
       #FB_STATE_TCP_RECONNECTING:
         REGION FB_STATE_TCP_RECONNECTING
           IF #tempTsendcStatus = #TSENDC_EST_OK THEN
             #statErrorAutoCleared := FALSE;
             //Monitor Connection
             #statFBState := #FB_STATE_OPERATING_MONITOR_TCP;
             // Begin MQTT Connection
             #statMqttConnectState := #MQTT_CONNECT_STATE_BUILD_PAKET;
           END_IF;
         END_REGION FB_STATE_TCP_RECONNECTING
       #FB_STATE_DISABLING: // Disabling active
         REGION DISABLING FB
           //  Disabling, e.g. closing connections, etc.
           // When disabling is complete the bit #statDisablingCompleted must be set
           // When MQTT is connected, send disconnect
           IF #statMqttConnectState = #MQTT_CONNECT_STATE_CONNECTED THEN
             IF #statTsendcReq = TRUE THEN
               //Interrupt any existing send jobs
               #statTsendcReq := FALSE;
             ELSE
               // INIT
               #statSendBufferPos := 0;
               //Build fixed Header
               //Message Type
               #statSendBuffer[#statSendBufferPos] := #MQTT_MSG_TYPE_DISCONNECT;
               #statSendBufferPos += 1;
               //Remaining Length (must be O)
               #statSendBuffer[#statSendBufferPos] := #REMAINIG_LEN_0;
               #statSendBufferPos += 1;
               //send request
               #statTsendcLen := #statSendBufferPos;
               #statTsendcReq := TRUE;
               #statMqttConnectState := #MQTT_CONNECT_STATE_DISCONNECTED;
             END_IF;
           ELSE
             //Disable TCP Connection
             #statTsendcReq := FALSE;
             #statTsendcEnable := FALSE;
             #statEnableTimerCommandWatchdog := TRUE;
           END_IF;
           // When TCP connection is closed
           IF #tempTsendcStatus = #TSENDC_DISCONNECTED THEN
             #statEnableTimerCommandWatchdog := FALSE;
             #statDisablingCompleted := TRUE;
           ELSIF #instTimerCommandWatchdog.Q THEN
             #statEnableTimerCommandWatchdog := FALSE;
             #statDisablingCompleted := TRUE;
           END_IF;
         END_REGION DISABLING FB
       ELSE // Undefined state in state machine reached
         #statStatus := #ERR_UNDEFINED_STATE;
         #statErrorUserCleared := TRUE;
     END_CASE;
   END_REGION STATE_MACHINE

   REGION OUTPUTS
     // Write outputs
     IF (#statDisablingCompleted = TRUE) THEN
       // Reset outputs if disabling completed
       #statValid := FALSE;
       #statBusy := FALSE;
       #statError := FALSE;
       #statDone := FALSE;
       #statErrorUserCleared := FALSE;
       #statErrorAutoCleared := FALSE;
       #statStatus := #STATUS_NO_CALL;
       // Reset application specific outputs
       #statRcvMsgStatus := #MSG_DECODE_STATUS_NO_NEW_MSG;
       #statRcvMsgDataLen := 0;
     ELSIF (#statErrorUserCleared = TRUE) AND (#statError = FALSE) THEN
       // Error can only be cleared by user; rising edge at enable input is needed to continue 
       #statValid := FALSE;
       #statBusy := FALSE;
       #statDone := FALSE;
       #statError := TRUE;
       // Write diagnostics
       #diagnostics.status := #statStatus;
       #diagnostics.subfunctionStatus := #statSubfunctionStatus;
       #diagnostics.stateNumber := #statFBErrorState;
       // execution aborted --> set state no processing
       #statTsendcEnable := FALSE; // Terminate Connection, no reason keep it up.
       #statFBState := #FB_STATE_NO_PROCESSING;
       #statMqttConnectState := #MQTT_CONNECT_STATE_NO_PROCESSING;
       #statMqttCommandState := #MQTT_COMMAND_STATE_NO_PROCESSING;
       #statRcvMsgDecodeState := #MSG_DECODE_STATE_NO_PROCESSING;

     ELSIF (#statErrorAutoCleared = TRUE) AND (#statError = FALSE) THEN
       // Error can be reset by FB automatically
       #statValid := FALSE;
       #statBusy := TRUE;
       #statError := TRUE;
       #statDone := FALSE;
       // Write diagnostics
       #diagnostics.status := #statStatus;
       #diagnostics.subfunctionStatus := #statSubfunctionStatus;
       #diagnostics.stateNumber := #statFBErrorState;
       // Handling of autocleared error
       CASE #statStatus OF
           //Just signal error and reset autocleared error afterwards.
         #ERR_MQTT_PAKET_ID_INVALID, #ERR_MQTT_SUBACK_FAILURE, #ERR_MQTT_CONNECT_TIMEOUT,
         #ERR_MQTT_COMMAND_SEND_TIMEOUT, #ERR_MQTT_COMMAND_MULTIPLE_INPUT, #ERR_CNT_EXCEEDS_ARRAY_DIMENSION,
         #ERR_MQTT_COMMAND_PUBLISH_TOPIC_INVALID, #ERR_QOS_INVALID, #ERR_MQTT_COMMAND_SUBSCRIBE_TOPIC_INVALID:
           #statErrorAutoCleared := FALSE;

         ELSE  // Statement section ELSE
           ;
       END_CASE;

     ELSIF (#statErrorAutoCleared = FALSE) AND (#statErrorUserCleared = FALSE) AND (#statError = TRUE) THEN
       // If autocleared error is acknowledged
       #statValid := TRUE;
       #statBusy := TRUE;
       #statError := FALSE;
       #statDone := FALSE;
       //   this line  more detailed status information is used instead of "#STATUS_SUBSEQUENT_CALL"
       CASE #statStatus OF
         #ERR_TCP_RECONNECTING, #ERR_MQTT_CONNECT_TIMEOUT:  // Reconnecting ok, start Mqtt reconnnect
           //set status
           #statStatus := #STATUS_MQTT_CONNECTING;
           //in the following status codes status stays connected. 
         #ERR_MQTT_PAKET_ID_INVALID, #ERR_MQTT_SUBACK_FAILURE, #ERR_MQTT_COMMAND_SEND_TIMEOUT,
         #ERR_MQTT_COMMAND_MULTIPLE_INPUT, #ERR_CNT_EXCEEDS_ARRAY_DIMENSION, #ERR_MQTT_COMMAND_PUBLISH_TOPIC_INVALID,
         #ERR_QOS_INVALID, #ERR_MQTT_COMMAND_SUBSCRIBE_TOPIC_INVALID:
           #statStatus := #STATUS_MQTT_CONNECTED;
         ELSE  // Statement section ELSE
           ;
       END_CASE;
     END_IF;

     // Write static values to outputs
     #valid := #statValid;
     #busy := #statBusy;
     #error := #statError;
     #status := #statStatus;
     //block sets ENO automatically:
     //ENO := TRUE;
     //Write application specific static values to outputs
     #done := #statDone;
     #receivedMsgStatus := #statRcvMsgStatus;
     #receivedMsgDataLen := #statRcvMsgDataLen;
   END_REGION OUTPUTS
END_FUNCTION_BLOCK

// folder: LMQTT/Utilities

FUNCTION "LMQTT_ConvertToUtf8" : Void   // FC6, SCL
TITLE = LMQTT_ConvertToUtf8
{ S7_Optimized_Access := 'TRUE' }
AUTHOR : SIEMENS
FAMILY : LMQTT
VERSION : 1.0
// Function to convert a WCHAR to a UTF-8 conformant byte sequence
   VAR_INPUT
      character : WChar;   // Character that shall be converted to UTF-8
   END_VAR
   VAR_OUTPUT
      convertedUtf8 : DWord;   // UTF-8 conformant byte sequence. B0 stores first Byte, B1 second and B2 third Byte. B3 is not used
      bytesUsed : USInt;   // Amount of Bytes converted. Ranges from 1 to 3.
      error : Bool;   // TRUE: An error occurred during the execution of the FC
      status : Word;   // 16#0000 - 16#7FFF: Status of the FC, 16#8000 - 16#FFFF: Error identification
   END_VAR
   VAR_TEMP
      tempStatus : Word;   // temp value for output 'status'
      tempConvertedUtf8 : DWord;   // temp value for output 'convertedUtf8'
      tempBytesUsed : USInt;   // temp value for output 'bytesUsed'
      tempCharacter : WChar;   // temp value for input 'character'
   END_VAR
   // Ret_Val : No return for this FC - see error and status output
   VAR CONSTANT
      STATUS_NO_ERROR : Word := 16#0000;   // no error status
      STATUS_EXECUTION_FINISHED : Word := 16#0000;   // Execution finished without errors
      ERR_UNDEFINED : Word := 16#8000;   // Error due to an undefined case
      USINT_NULL : USInt := 0;   // Init value with 0
      DWORD_NULL : DWord := 16#0000_0000;   // Init value with 0
      EMPTY_WCHAR : WChar := WCHAR#' ';   // Empty WChar for comparison
      BELOW_7F : Word := 16#007F;   // Upper limit for character if only one Byte used
      BELOW_7FF : Word := 16#07FF;   // Upper limit for character if two Byte used
      BELOW_MAX_FFFF : Word := 16#FFFF;   // Upper limit for character if three Byte used
      BYTE_3F : Byte := 16#3F;   // Conversion Value
      BYTE_80 : Byte := 16#80;   // Conversion Value
      BYTE_C0 : Byte := 16#C0;   // Conversion Value
      BYTE_E0 : Byte := 16#E0;   // Conversion Value
      USINT_ONE : USInt := 1;   // Const Value to assign amount of bytes used
      USINT_TWO : USInt := 2;   // Const Value to assign amount of bytes used
      USINT_THREE : USInt := 3;   // Const Value to assign amount of bytes used
   END_VAR
BEGIN
   REGION BLOCK INFO HEADER
       //=============================================================================
       // SIEMENS AG
       // (c)Copyright 2020
       //-----------------------------------------------------------------------------
       // Library:       LMQTT
       // Tested with:   CPU 1516-3 PN/DP V2.8
       // Engineering:   TIA Portal V16
       // Restrictions:  --
       // Requirements:  --
       // Functionality: Converts a single WChar Character to a valid UTF-8 encoded byte sequence and saves this to a DWord.
       //                The amount of bytes saved is stored in bytesUsed Output.
       //-----------------------------------------------------------------------------
       // Change log table:
       // Version    Date         Expert in charge         Changes applied
       // 03.00.00   01.10.2020   Siemens Online Support   First released version
       //=============================================================================
   END_REGION

   REGION INITIALISATION  
       // Initialize functionality: reset of variables, diagnostics, etc.
       #tempConvertedUtf8 := #DWORD_NULL;
       #tempBytesUsed := #USINT_NULL;
       #tempStatus := #STATUS_NO_ERROR;
       //assign temp value from input:
        #tempCharacter := #character;

   END_REGION

   REGION PROGRAM LOGIC
       // Use this region for application specific code
       IF #tempCharacter = #EMPTY_WCHAR THEN
           //will be only 1 byte occupied
           #tempConvertedUtf8 := WCHAR_TO_DWORD(#tempCharacter);
           #tempBytesUsed := #USINT_ONE;
       ELSIF (WCHAR_TO_WORD(#tempCharacter) <= (#BELOW_7F)) THEN
           //will be only 1 byte occupied
           #tempConvertedUtf8 := WCHAR_TO_DWORD(#tempCharacter);
           #tempBytesUsed := #USINT_ONE;
       ELSIF (WCHAR_TO_WORD(#tempCharacter) <= (#BELOW_7FF)) THEN
           //will be 2 byte occupied
           #tempConvertedUtf8.%B1 := (WCHAR_TO_BYTE(#tempCharacter) AND #BYTE_3F) OR #BYTE_80;
           #tempConvertedUtf8.%B0 := WORD_TO_BYTE(SHR(IN := WCHAR_TO_WORD(#tempCharacter), N := 6)) OR #BYTE_C0;
           #tempBytesUsed := #USINT_TWO;
       ELSIF (WCHAR_TO_WORD(#tempCharacter) <= (#BELOW_MAX_FFFF)) THEN
           //will be 3 byte occupied
           #tempConvertedUtf8.%B2 := (WCHAR_TO_BYTE(#tempCharacter) AND #BYTE_3F) OR #BYTE_80;
           #tempConvertedUtf8.%B1 := (WORD_TO_BYTE(SHR(IN := WCHAR_TO_WORD(#tempCharacter), N := 6)) AND #BYTE_3F) OR #BYTE_80;
           #tempConvertedUtf8.%B0 := WORD_TO_BYTE(SHR(IN := WCHAR_TO_WORD(#tempCharacter), N := 12)) OR #BYTE_E0;
           #tempBytesUsed := #USINT_THREE;
       END_IF;
   END_REGION

   REGION OUTPUTS
       // Write application specific temp values to outputs
       #bytesUsed := #tempBytesUsed;
       #convertedUtf8 := #tempConvertedUtf8;
       // Write error and status
       #error := #tempStatus.%X15;
       #status := #tempStatus;
       // ENO mechanism is not used --> ENO := TRUE;
       ENO := TRUE;
   END_REGION
END_FUNCTION

// folder: LStream

FUNCTION_BLOCK "LStream_JsonDeserializer"   // FB3, SCL
TITLE = LStream_JsonDeserializer / LStream_JsonParser
{ S7_Optimized_Access := 'TRUE' }
AUTHOR : DI_FA_S_SUP_EuC
FAMILY : LStream
VERSION : 1.0
// parses a JSON string provided in the raw paramter  and rebuilds the coinatend bytes into a tree structure / Parses JSON file, with or without seach option
   VAR_INPUT
      execute : Bool;   // Rising edge starts action once
      search : Bool;   // TRUE: Search option is acticve
   END_VAR
   VAR_OUTPUT
      done : Bool;   // TRUE: Commanded functionality has been completed successfully
      busy : Bool;   // TRUE: FB is not finished and new output values can be expected
      error : Bool;   // TRUE: An error occurred during the execution of the FB
      status : Word := 16#7000;   // 16#0000 - 16#7FFF: Status of the FB, 16#8000 - 16#FFFF: Error identification
      resultCount : Int;   // Count of parsed JSON elements
   END_VAR
   VAR_IN_OUT
      tree : Array[*] of "LStream_typeElement";   // JSON tree containing the stored data
      raw : Array[*] of Byte;   // raw JSON data to parse in byte format
   END_VAR
   VAR
      statExecuteOld : Bool;   // Old value of 'execute' input for edge detection
      statDone : Bool;   // Static value for output 'done'
      statBusy : Bool;   // Static value for output 'busy'
      statError : Bool;   // Static value for output 'error'
      statStatus : Word := 16#7000;   // Static value for output 'status'
      statFBState : DInt := 0;   // State in the state machine of the FB
      statCountOfTree : Int;   // Static count of tree fields
      statCountOfRaw : Int;   // Static count of raw fields
      statResultCount : Int;   // Static value of result count
      statRawIndex : Int;   // Static value of raw index
      instWatchdog : IEC_TIMER;   // instance of watchdog timer
      statSearch : Bool;   // TRUE: Only keys provided in tree will be parsed
      statKeyValueFound : Bool;   // TRUE: Key exisits in raw data
      statTreeIndex : Int;   // Static value of tree index
      statSearchIndex : DInt;   // Static search
      statDepth : SInt := -1;   // Static value of JSON depth
      statOpen : Bool;   // TRUE: Key or Value is opened
      statInfoStartIndex : Int;   // Start index of current info in raw key or value
      statIgnorableCharacter : Bool;   // Next character to be ignored
      statInfoLen : UInt;   // Current information length key or value
      statKey : String;   // Static key string
      statValue : String;   // Static value string
      statKeyNotFoundCount : Int;   // Count of provided keys that weren't found
      statArrayOpen : Bool;   // TRUE: New JSON array is open
      statObjectArray : Bool;   // TRUE: Is type array of obejct
      statType : SInt;   // Current type of element
      statDefineValueType : Bool;   // TRUE: Value Type can be defined
      statArrayName : String;   // Name of array
   END_VAR
   VAR_TEMP
      tempExecute : Bool;   // Temporary value for input 'execute'
      tempRawIndex : Int;   // Index of raw field
      tempKeyToFind : String;   // Provided key to which the value should be found
      tempSearchResult : DInt;   // Temp value of search result
   END_VAR
   VAR CONSTANT
      FB_STATE_NO_PROCESSING : DInt := 0;   // FB state: No processing
      FB_STATE_PARSE : DInt := 1;   // FB state: Processing Parsing
      STATUS_EXECUTION_FINISHED : Word := 16#0000;   // Execution finished without errors
      STATUS_NO_CALL : Word := 16#7000;   // No job being currently processed
      STATUS_FIRST_CALL : Word := 16#7001;   // First call after incoming new job (rising edge 'execute')
      STATUS_SUBSEQUENT_CALL : Word := 16#7002;   // Subsequent call during active processing without further details
      ERR_TREE_ARRAY_TOO_SMALL : Word := 16#8201;   // Error: provided array to too small
      ERR_EMPTY_RAW_DATA : Word := 16#8401;   // Error: no raw data provided
      ERR_UNDEFINED_STATE : Word := 16#8600;   // Error: due to an undefined state in state machine
      JSON_QUTATIONMARK : Byte := 16#22;   // ASCII code for '"'
      JSON_COLON : Byte := 16#3A;   // ASCII code for ':'
      JSON_COMMA : Byte := 16#2C;   // ASCII code for ','
      JSON_BRACES_OPEN : Byte := 16#7B;   // ASCII code for '{'
      JSON_BRACES_CLOSE : Byte := 16#7D;   // ASCII code for '}'
      JSON_BRACKETS_OPEN : Byte := 16#5B;   // ASCII code for '['
      JSON_BRACKETS_CLOSE : Byte := 16#5D;   // ASCII code for ]
      "JSON_PROTECTION_KEY_\" : Byte := 16#5C;   // ASCII coder for / indicates closing / ASCII coder for \ indicates closing
      "JSON_CLOSE_KEY_/" : Byte := 16#2F;   // ASCII coder for / indicates closing
      LINE_FEED : Byte := 16#0A;   // ASCII code for line feed
      TAB : Byte := 16#09;   // ASCII code for TAB
      CARRIAGE_RETURN : Byte := 16#0D;   // ASCII code for carriage return
      SPACE : Byte := 16#20;   // ASCII code for blank space
      FIRST_DIM : USInt := 1;   // Constant for first array dimension
      MAX_LOOP_TIME : Time := T#3ms;   // Max duration of loop, will be continued in next cycle
      INVALID_SEARCH : DInt := -1;   // Return value if Search in LParse_FindStringInCharrArrayAdv was not successfull
      KEY_NOT_FOUND : String := 'Key not found';   // Value string in case key wasn't found
      INCREMENT_BY_ONE : USInt := 1;   // Constant to increment by one
      DECREMENT_BY_ONE : SInt := 1;   // Constant to decrement by one
      DECREMENT_BY_TWO : SInt := 2;   // Constant to decrement by one / Constant to decrement by two
      OBJECT : SInt := 0;   // Constant for value typ object / Constant for typ object
      "ARRAY" : SInt := 1;   // Constant for value typ array / Constant for typ array
      "STRING" : SInt := 2;   // Constant for value type string
      NUMBER : SInt := 3;   // Constant for value type number
      BOOLEAN : SInt := 4;   // Constant for value type boolean
      DEPTH_NOT_DEFINED : Int := -1;   // Constant indicating depth wasn't yet defined
   END_VAR
BEGIN
   REGION BLOCK INFO HEADER
     //===============================================================================
     // SIEMENS AG / (c)Copyright 2021
     //-------------------------------------------------------------------------------
     // Title:            LStream_JsonDeserializer
     // Comment/Function: parses a JSON string provided in the raw paramter
     //                   and rebuilds the coinatend bytes into a tree structure
     // Library/Family:   LStream
     // Author:           DI FA S SUP E&C
     // Tested with:      S7-1500 V2.8
     // Engineering:      TIA Portal V16
     // Restrictions:     -- 
     // Requirements:     LStream_FindStringInByteArrayAdv(FC), LStream_typeElement(UDT)
     //-------------------------------------------------------------------------------
     // Change log table:
     // Version  | Date       | Expert in charge       | Changes applied
     //----------|------------|------------------------|------------------------------
     // 01.0.0 | 2021-03-10 | DI FA S SUP E&C          | First released version
     // 01.0.8 | 2021-09-23 | DI FA S SUP E&C          | Adjustment type definition & bug fixes
     //===============================================================================
   END_REGION

   #tempExecute := #execute; // Work with temporary value / create process image

   REGION TRIGGERING
     IF (#tempExecute = TRUE) AND (#statExecuteOld = FALSE) // Check if FB is triggered
       AND (#statStatus = #STATUS_NO_CALL)
     THEN // First call; initialize FB
       #statDone := FALSE;
       #statBusy := TRUE;
       #statError := FALSE;
       #statStatus := #STATUS_FIRST_CALL;
       // State machine - start processing
       #statFBState := #FB_STATE_PARSE;

       // Initialize functionality: reset of variables, diagnostics, etc.
       #statSearch := #search;
       #statCountOfRaw := DINT_TO_INT(UPPER_BOUND(ARR := #raw, DIM := #FIRST_DIM));
       #statCountOfTree := DINT_TO_INT(UPPER_BOUND(ARR := #tree, DIM := #FIRST_DIM));
       #statOpen := FALSE;
       #statDepth := -1;
       #statRawIndex := 0;
       #statTreeIndex := 0;
       #statInfoLen := 0;
       #statSearchIndex := 0;
       #statKeyNotFoundCount := 0;
       #statType := -1;
       #statDefineValueType := FALSE;
       #statObjectArray := FALSE;

     ELSIF (#statStatus = #STATUS_FIRST_CALL) THEN
       #statStatus := #STATUS_SUBSEQUENT_CALL;
     END_IF;

     // Edge detection 'execute' input
     #statExecuteOld := #tempExecute;
   END_REGION TRIGGERING

   IF (#statStatus = #STATUS_NO_CALL) THEN // Nothing to do -> End here to reduce "system load"
     RETURN;
   END_IF;

   REGION STATE_MACHINE

     CASE #statFBState OF // State machine of FB
       #FB_STATE_NO_PROCESSING:
         REGION NO PROCESSING
           // No processing active (Note: this state must always be present and left empty)
           ;
         END_REGION NO PROCESSING

       #FB_STATE_PARSE: // Processing active
         REGION PARSING

           //rest watchdog
           #instWatchdog.TON(IN := FALSE,
                             PT := #MAX_LOOP_TIME);
           //start watchdog
           #instWatchdog.TON(IN := TRUE,
                             PT := #MAX_LOOP_TIME);

           FOR #tempRawIndex := #statRawIndex TO #statCountOfRaw DO

             REGION FIND KEY
               //pre check if key exist in raw data, if search option is active
               IF (#statSearch AND #statKeyValueFound = FALSE) THEN
                 IF (#statTreeIndex < #statCountOfTree) THEN
                   #tempSearchResult := "LStream_FindStringInByteCharArrayAdv"(searchFor := #tree[#statTreeIndex].key, startPosition := #statSearchIndex, searchIn := #raw);
                   IF (#tempSearchResult = #INVALID_SEARCH) THEN
                     //case key not found
                     #tree[#statTreeIndex].value := #KEY_NOT_FOUND;
                     #statTreeIndex += #INCREMENT_BY_ONE;
                     #statKeyNotFoundCount += #INCREMENT_BY_ONE;
                   ELSE//case key found
                     //move read pointer to last found index
                     #statSearchIndex := #tempSearchResult;
                     #statKeyValueFound := TRUE;
                   END_IF;
                 END_IF;
               END_IF;
             END_REGION FIND KEY   


             CASE #raw[#tempRawIndex] OF

               #JSON_BRACES_OPEN:
                 REGION OBJECT OPEN     

                   #statDepth += USINT_TO_SINT(#INCREMENT_BY_ONE);
                   IF (#statDefineValueType) THEN
                     #statDefineValueType := FALSE;
                     #statType := #OBJECT;
                     #tree[#statTreeIndex - #DECREMENT_BY_ONE].type := #statType;
                   END_IF;
                 END_REGION OBJECT OPEN

               #JSON_BRACES_CLOSE:
                 REGION OBJECT CLOSE      

                   #statDepth -= #DECREMENT_BY_ONE;
                   //last element closed, and there is still info in the buffer, then write value to last key
                   IF (#statDepth = -1 AND #statInfoLen > 0) THEN
                     //in case of 0 length, Chars_To_Strig returns the maxium possible char combination
                     Chars_TO_Strg(Chars := #raw,
                                   pChars := #statInfoStartIndex,
                                   Cnt := #statInfoLen,
                                   Strg => #statValue);
                     #statInfoLen := 0;

                     //value Type wasn't yet definied must be either number or boolean
                     IF (#statDefineValueType) THEN
                       #statDefineValueType := FALSE;

                       IF #statValue = 'FALSE' OR #statValue = 'TRUE'
                         OR #statValue = 'false' OR #statValue = 'true' THEN
                         #statType := #BOOLEAN;
                       ELSE
                         #statType := #NUMBER;
                       END_IF;

                     END_IF;

                     IF (#statSearch) THEN

                       IF (#statTreeIndex > 0) THEN
                         //in case of 0 length, Chars_To_Strig returns the maxium possible char combination
                         IF (#statKey = #tree[#statTreeIndex - #DECREMENT_BY_ONE].key) THEN
                           //only write into tree, if key matches, otherwise continue with search for matching key
                           #tree[#statTreeIndex - #DECREMENT_BY_ONE].value := #statValue;
                           #tree[#statTreeIndex - #DECREMENT_BY_ONE].type := #statType;
                           #statKeyValueFound := FALSE;
                         END_IF;
                       ELSE 
                         IF (#statKey = #tree[#statTreeIndex].key) THEN
                           #tree[#statTreeIndex].value := #statValue;
                           #tree[#statTreeIndex].type := #statType;
                           #statKeyValueFound := FALSE;
                         END_IF;
                       END_IF;

                     ELSE // IF #search option isn't active (parse all) add key TO the current #tree index
                       #tree[#statTreeIndex - #DECREMENT_BY_ONE].value := #statValue;
                       #tree[#statTreeIndex - #DECREMENT_BY_ONE].type := #statType;
                     END_IF;
                   END_IF;
                 END_REGION OBJECT CLOSE

               #JSON_BRACKETS_OPEN:
                 REGION ARRAY OPEN

                   #statDepth += USINT_TO_SINT(#INCREMENT_BY_ONE);

                   IF (#statTreeIndex > 0) THEN
                     //
                     #tree[#statTreeIndex - #DECREMENT_BY_ONE].type := #ARRAY;

                     //save arrayName
                     #statArrayName := #tree[#statTreeIndex - #DECREMENT_BY_ONE].key;

                     #statTreeIndex += #INCREMENT_BY_ONE;

                   ELSE // first element, is of type array
                     #tree[#statTreeIndex].type := #ARRAY;
                   END_IF;

                   #statArrayOpen := TRUE;
                   #statObjectArray := FALSE;
                 END_REGION ARRAY OPEN

               #JSON_BRACKETS_CLOSE:
                 REGION ARRAY CLOSE
                   #statDepth -= #DECREMENT_BY_ONE;
                   #statArrayOpen := FALSE;

                 END_REGION ARRAY CLOSE

               #JSON_QUTATIONMARK:
                 REGION QUTATIONMARK
                   IF (#statOpen) THEN
                     IF (NOT (#raw[#tempRawIndex - #DECREMENT_BY_ONE] = #"JSON_PROTECTION_KEY_\")) THEN
                       // previous sign \ then allowed in string adjust
                       #statOpen := FALSE;
                     ELSE
                       #statInfoLen += #INCREMENT_BY_ONE;
                     END_IF;
                   ELSE
                     #statInfoStartIndex := #tempRawIndex + #INCREMENT_BY_ONE; //set reader to next sign
                     #statOpen := TRUE;
                     #statIgnorableCharacter := FALSE;
                     //Qutation mark after colomn indicates value is of type string
                     IF #statDefineValueType THEN
                       #statType := #STRING;
                       #tree[#statTreeIndex - #DECREMENT_BY_ONE].type := #statType;
                       #statDefineValueType := FALSE;
                     END_IF;

                   END_IF;
                 END_REGION QUTATIONMARK

               #JSON_COLON:
                 REGION COLON

                   //array is open, and a sperate key is found indication for array of objects
                   //
                   IF #statArrayOpen AND NOT #statObjectArray THEN
                     #statObjectArray := TRUE;
                     #statTreeIndex -= #DECREMENT_BY_ONE;
                   END_IF;

                   //error handling
                   IF (#statTreeIndex > #statCountOfTree) THEN
                     //data does not fit in the provided tree 
                     #statStatus := #ERR_TREE_ARRAY_TOO_SMALL;
                     #statDone := TRUE;
                     EXIT;
                   END_IF;

                   //write key, if colon is part of a string
                   IF (NOT #statOpen) THEN
                     Chars_TO_Strg(Chars := #raw,
                                   pChars := #statInfoStartIndex,
                                   Cnt := #statInfoLen,
                                   Strg => #statKey);
                     #statInfoLen := 0;

                     //After key was written, type of value can be definied, value can be object, array, string, number, or boolean
                     #statDefineValueType := TRUE;

                     IF (#statSearch) THEN
                       //only write into tree, if key matches, otherwise continue with search for matching key
                       IF (#statKey = #tree[#statTreeIndex].key) THEN
                         //#tree[#statTreeIndex].type := #statType;
                         #tree[#statTreeIndex].depth := #statDepth;
                         #statTreeIndex += #INCREMENT_BY_ONE;
                       END_IF;

                     ELSE// if search option isn't active (parse all) the add key to the current tree index 
                       #tree[#statTreeIndex].key := #statKey;
                       //#tree[#statTreeIndex].type := #statType;
                       #tree[#statTreeIndex].depth := #statDepth;
                       #tree[#statTreeIndex].value := 'NULL';
                       #statTreeIndex += #INCREMENT_BY_ONE;
                     END_IF;

                     #statInfoStartIndex := #tempRawIndex+1;

                   ELSE//case : included in string
                     #statInfoLen += #INCREMENT_BY_ONE;
                   END_IF;
                 END_REGION COLON

               #JSON_COMMA:
                 REGION COMMA

                   //error handling
                   IF (#statTreeIndex > #statCountOfTree + #INCREMENT_BY_ONE) THEN
                     //data does not fit in the provided tree 
                     #statStatus := #ERR_TREE_ARRAY_TOO_SMALL;
                     #statDone := TRUE;
                     EXIT;
                   END_IF;

                   IF (NOT #statOpen) THEN
                     //write value comma isn't part of string
                     IF (#statInfoLen > 0) THEN
                       //in case of 0 length, Chars_To_Strig returns the maxium possible char combination
                       Chars_TO_Strg(Chars := #raw,
                                     pChars := #statInfoStartIndex,
                                     Cnt := #statInfoLen,
                                     Strg => #statValue);
                       #statInfoLen := 0;
                     ELSE
                       #statValue := 'NULL';
                       #statDefineValueType := FALSE;
                       //no value Type deafult value type NULL/Default is correct
                     END_IF;

                     //value Type wasn't yet definied must be either number or boolean
                     IF (#statDefineValueType) THEN
                       #statDefineValueType := FALSE;

                       IF #statValue = 'FALSE' OR #statValue = 'TRUE'
                         OR #statValue = 'false' OR #statValue = 'true' THEN
                         #statType := #BOOLEAN;
                       ELSE
                         #statType := #NUMBER;
                       END_IF;

                     END_IF;
                     //add value always to the last JSON element
                     IF (#statSearch) THEN

                       IF (#statTreeIndex > 0) THEN
                         //in case of 0 length, Chars_To_Strig returns the maxium possible char combination
                         IF (#statKey = #tree[#statTreeIndex - #DECREMENT_BY_ONE].key) THEN
                           //only write into tree, if key matches, otherwise continue with search for matching key
                           #tree[#statTreeIndex - #DECREMENT_BY_ONE].value := #statValue;
                           #tree[#statTreeIndex].type := #statType;
                           #statKeyValueFound := FALSE;
                         END_IF;
                       ELSE
                         IF (#statKey = #tree[#statTreeIndex].key) THEN
                           // if search option isn't active (parse all) the add key to the current tree index 
                           #tree[#statTreeIndex].value := #statValue;
                           #tree[#statTreeIndex].type := #statType;
                           #statKeyValueFound := FALSE;
                         END_IF;
                       END_IF;

                     ELSE//search option isn't active
                       #tree[#statTreeIndex - #DECREMENT_BY_ONE].value := #statValue;
                       #tree[#statTreeIndex - #DECREMENT_BY_ONE].type := #statType;
                       //case simple array last information
                       IF (#tree[#statTreeIndex - #DECREMENT_BY_ONE].depth = #DEPTH_NOT_DEFINED) THEN
                         #tree[#statTreeIndex - #DECREMENT_BY_ONE].depth := #tree[#statTreeIndex - #DECREMENT_BY_TWO].depth;
                         #tree[#statTreeIndex - #DECREMENT_BY_ONE].key := #statArrayName;
                         //always take depth from previous entry of simple array e.g "ArrayName":["ArrayValue1","ArrayValue2"]
                       END_IF;
                     END_IF;

                     IF (#statArrayOpen AND NOT #statObjectArray) THEN
                       //only write if Array is open and simple array
                       //
                       #tree[#statTreeIndex- #DECREMENT_BY_ONE].key := #statArrayName;
                       #tree[#statTreeIndex - #DECREMENT_BY_ONE].depth := #statDepth;//#tree[#statTreeIndex - #DECREMENT_BY_TWO].depth +1;
                       #tree[#statTreeIndex- #DECREMENT_BY_ONE].type := #statType;
                       //always take depth from previous entry of simple array e.g "ArrayName":["ArrayValue1","ArrayValue2"]


                       // #tree[#statTreeIndex].key := #tree[#statTreeIndex - #DECREMENT_BY_ONE].key;
                       // #tree[#statTreeIndex].depth := #tree[#statTreeIndex - #DECREMENT_BY_ONE].depth;
                       // #tree[#statTreeIndex].type := #tree[#statTreeIndex - #DECREMENT_BY_ONE].type;
                       #statTreeIndex += #INCREMENT_BY_ONE;
                     END_IF;

                     #statInfoStartIndex := #tempRawIndex;

                   ELSE//case ; included in string
                     #statInfoLen += #INCREMENT_BY_ONE;
                   END_IF;
                 END_REGION

               #TAB, #LINE_FEED, #CARRIAGE_RETURN, #SPACE:
                 REGION READ TAB LINE FEED CARRIAGE RETURN   
                   IF (NOT #statOpen) THEN
                     //do nothing when tab, line feed, or carriage return
                     #statIgnorableCharacter := TRUE;
                   ELSE//case space included in string
                     #statInfoLen += #INCREMENT_BY_ONE;
                   END_IF;

                 END_REGION READ TAB LINE FEED CARRIAGE RETURN     


               ELSE // all other characters
                 REGION ALL OTHER SIGNS
                 IF (#statIgnorableCharacter = TRUE) THEN
                   #statIgnorableCharacter := FALSE;
                   #statInfoStartIndex := #tempRawIndex; // set KeyIndex after all ignorableCharacters are read
                   #statInfoLen += #INCREMENT_BY_ONE;
                 ELSE
                   #statInfoLen += #INCREMENT_BY_ONE;
                 END_IF;
                 END_REGION ALL OTHER SIGNS 
             END_CASE;

             #statRawIndex := #tempRawIndex;

             //quit and resume in next cycle if watchdogtimer is exceed
             IF (#instWatchdog.Q) THEN
               #statRawIndex += #INCREMENT_BY_ONE;
               EXIT;
             END_IF;

           END_FOR;

           //if parser is through the entire raw data or end of tree array reached
           IF (#statRawIndex >= #statCountOfRaw) OR (#statTreeIndex > #statCountOfTree) THEN
             #statStatus := #STATUS_EXECUTION_FINISHED;
             #statResultCount := #statTreeIndex - #statKeyNotFoundCount;
           END_IF;
         END_REGION PARSING

       ELSE // Undefined state in state machine reached
         REGION UNDEFINED STATE
           #statStatus := #ERR_UNDEFINED_STATE;
         END_REGION UNDEFINED STATE
     END_CASE;
   END_REGION STATE_MACHINE

   REGION OUTPUTS
     // Write outputs
     IF (#statStatus = #STATUS_EXECUTION_FINISHED) AND (#statDone = FALSE) THEN // Execution finished without errors
       REGION EXECUTION FINSIHED
         #statDone := TRUE;
         #statBusy := FALSE;
         #statError := FALSE;
         // execution aborted --> set state no processing
         #statFBState := #FB_STATE_NO_PROCESSING;
       END_REGION EXECUTION FINSIHED

     ELSIF (#statStatus.%X15 = TRUE) AND (#statError = FALSE) THEN // Error occurred (#statStatus is 16#8000 to 16#FFFF)
       REGION ERROR OCCURD
         #statDone := FALSE;
         #statBusy := FALSE;
         #statError := TRUE;
         // execution aborted --> set state no processing
         #statFBState := #FB_STATE_NO_PROCESSING;
       END_REGION ERROR OCCURD

     ELSIF (#tempExecute = FALSE) AND ((#statDone = TRUE) OR (#statError = TRUE)) THEN // Reset outputs
       REGION EXECUTE RESETED
         #statDone := FALSE;
         #statBusy := FALSE;
         #statError := FALSE;
         #statStatus := #STATUS_NO_CALL;
         // Reset application specific outputs
         #statResultCount := 0;
       END_REGION EXECUTE RESETED
     END_IF;

     REGION WRITE STATIC VALUES TO OUTPUTS
       #done := #statDone;
       #busy := #statBusy;
       #error := #statError;
       #status := #statStatus;

       ENO := TRUE;
       // Write application specific static values to outputs
       #resultCount := #statResultCount;
     END_REGION WRITE STATIC VALUES TO OUTPUT
   END_REGION OUTPUTS
END_FUNCTION_BLOCK

FUNCTION_BLOCK "LStream_JsonSerializer"   // FB5, SCL
TITLE = LStream_JsonDeserializer / LStream_JsonParser
{ S7_Optimized_Access := 'TRUE' }
AUTHOR : DI_FA_S_SUP_EuC
FAMILY : LStream
VERSION : 1.0
// parses a JSON string provided in the raw paramter  and rebuilds the coinatend bytes into a tree structure / Parses JSON file, with or without seach option
   VAR_INPUT
      execute : Bool;   // Rising edge starts action once
   END_VAR
   VAR_OUTPUT
      done : Bool;   // TRUE: Commanded functionality has been completed successfully
      busy : Bool;   // TRUE: FB is not finished and new output values can be expected
      error : Bool;   // TRUE: An error occurred during the execution of the FB
      status : Word := 16#7000;   // 16#0000 - 16#7FFF: Status of the FB, 16#8000 - 16#FFFF: Error identification
      count : UInt;   // Count of char/ byte info elements in byte array / Count of parsed JSON elements
   END_VAR
   VAR_IN_OUT
      tree : Array[*] of "LStream_typeElement";   // JSON tree containing the stored data
      jsonByteArray : Array[*] of Byte;   // JSON structure as array of bytes / raw JSON data to parse in byte format
   END_VAR
   VAR
      statExecuteOld : Bool := FALSE;   // Old value of 'execute' input for edge detection
      statDone : Bool := FALSE;   // Static value for output 'done'
      statBusy : Bool := FALSE;   // Static value for output 'busy'
      statError : Bool := FALSE;   // Static value for output 'error'
      statCount : UInt := 0;   // Static value for ouput 'count'
      statStatus : Word := 16#7000;   // Static value for output 'status'
      statFbState : DInt := 0;   // State in the state machine of the FB
      statFbPreviousState : DInt := 0;   // Previos state in the state machine of the FB
      statFbNextState : DInt := 0;   // Next state in the state machine of the FB
      statIndexJsonByteArray : UInt := 0;   // Index indicating current element of byte array to be written
      statIndexTreeArray : UInt := 0;   // Index indicating current element of tree array to be read
      statTreeLen : DInt := 0;   // Length of tree array
      statJsonByteLen : DInt := 0;   // Length of xml byte array / Length of json byte array
      statInfoToWrite : String := '';   // Static value of current information that should be written to XML
      statIsLastElement : Bool := FALSE;   // TRUE: is last element in tree array
      statLastElementIsClosed : Bool := FALSE;   // TRUE: Last JSON element is closed / TRUE: Last XML element is closed
      statStackIndexOpenElement : Array[0..#STACK_SIZE] of Char;   // Stack of open elements
      statStackIndex : Int := -1;   // Stack pointer and current depth / Stack pointer
      instWatchdog : IEC_TIMER;   // Instance for watchdog timer
      statIsArrayOpen : Bool;   // Static value indicating weather an array is open
      statIsArrayFieldClosed : Bool;   // Static value indicating weather an array field was closed
      statIsFirstElement : Bool;   // TRUE: first field of simple array
      statFirstArrayKey : String;   // First key of array, used to check for new array beginning
      statArrayName : String;   // Name of Array
   END_VAR
   VAR_TEMP
      tempExecute : Bool;   // Temporary value for input 'execute'
      tempCntCharsAdded : UInt;   // Temporary value indicating count of chars added to byte array
   END_VAR
   VAR CONSTANT
      FB_STATE_NO_PROCESSING : DInt := 0;   // FB state: No processing
      FB_STATE_NEXT_ELEMENT : DInt := 1;   // FB state: Get Next Element
      FB_STATE_VALUE_TYPE : DInt := 2;   // FB state: Switch Value type / FB state: Switch Element type
      FB_STATE_WRITE_TO_JSON : DInt := 3;   // FB state: Add Informationto xml byte array
      FB_STATE_CLOSE_STACK_ELEMENT : DInt := 4;   // FB state: Close Parent Element
      STATUS_EXECUTION_FINISHED : Word := 16#0000;   // Execution finished without errors
      STATUS_NO_CALL : Word := 16#7000;   // No job being currently processed
      STATUS_FIRST_CALL : Word := 16#7001;   // First call after incoming new job (rising edge 'execute')
      STATUS_SUBSEQUENT_CALL : Word := 16#7002;   // Subsequent call during active processing without further details
      ERR_UNDEFINED_STATE : Word := 16#8600;   // Error: due to an undefined state in state machine
      ERR_IN_BLOCK_OPERATION : Word := 16#8001;   // Error: wrong operation of the function block
      ERR_PARAMETRIZATION : Word := 16#8200;   // Error: during parameterization
      ERR_PROCESSING_EXTERN : Word := 16#8400;   // Error: when processing from outside (e. g. wrong I/O signals, axis not referenced)
      ERR_UNDEFINED_TYPE : Word := 16#8401;   // Error: user enter undefined type
      ERR_UNEXPECTED_DEPTH : Word := 16#8402;   // Error: provided json tree structure is too deep / Error: provided xml tree structure is too deep
      ERR_DEPTH_MISSING : Word := 16#8403;   // Error: provided json tree structure does not contain correct depth / Error: provided xml tree structure does not contain correct depth
      ERR_PROCESSING_INTERN : Word := 16#8600;   // Error: when processing internally (e. g. when calling a system function)
      ERR_TREE_OUT_OF_BOUNDS : Word := 16#8601;   // Error: tree array out of bounds
      ERR_JSON_OUT_OF_BOUNDS : Word := 16#8602;   // Error: byte array out of bounds
      ERR_STACK_OUT_OF_BOUNDS : Word := 16#8603;   // Error: stack array out of bounds
      ERR_AREA_RESERVED : Word := 16#8800;   // Error: reserved area
      ERR_USER_DEFINED_CLASSES : Word := 16#9000;   // Error: user-defined error classes
      QUTATIONMARK : Char := '"';   // ASCII code for '"'
      COLON : Char := ':';   // ASCII code for ':'
      COMMA : Char := ',';   // ASCII code for ','
      BRACES_OPEN : Char := '{';   // ASCII code for '{'
      BRACES_CLOSE : Char := '}';   // ASCII code for '}'
      BRACKETS_OPEN : Char := '[';   // ASCII code for '['
      BRACKETS_CLOSE : Char := ']';   // ASCII code for ]
      "PROTECTION_KEY_\" : Char := '\';   // ASCII coder for / indicates closing / ASCII coder for \ indicates closing
      LINE_FEED : Char := '$L';   // ASCII code for line feed
      TAB : Char := '$T';   // ASCII code for TAB
      CARRIAGE_RETURN : Char := '$R';   // ASCII code for carriage return
      SPACE : Char := ' ';   // ASCII code for blank space
      FIRST_DIM : USInt := 1;   // Constant for first array dimension
      MAX_REPEAT_TIME : Time := T#3ms;   // Max duration of loop, will be continued in next cycle
      INVALID_SEARCH : DInt := -1;   // Return value if Search in LParse_FindStringInCharrArrayAdv was not successfull
      KEY_NOT_FOUND : String := 'Key not found';   // Value string in case key wasn't found
      INCREMENT_BY_ONE : USInt := 1;   // Constant to increment by one
      DECREMENT_BY_ONE : SInt := 1;   // Constant to decrement by one
      OBJECT : SInt := 0;   // Constant for value typ object / Constant for typ object
      "ARRAY" : SInt := 1;   // Constant for value typ array / Constant for typ array
      "STRING" : SInt := 2;   // Constant for value type string
      NUMBER : SInt := 3;   // Constant for value type number
      BOOLEAN : SInt := 4;   // Constant for value type boolean
      NEXT_INDEX : UInt := 1;   // Constant value to get next index
      STACK_SIZE : UInt := 10;   // Constant for Stack Size, equals max depth
      WHITE_SPACE : Char := ' ';   // ASCII code for white space
      NOT_INITALYZED : SInt := -1;   // Constant value representing not initalyzed tree element
      EMPTY : String;   // Constant value representing an empty string
      NULL : String := 'NULL';   // Constant value representing null
   END_VAR
   // statStackIndexOpenElement[0] := '$00';
   // statStackIndexOpenElement[1] := '$00';
BEGIN
   REGION BLOCK INFO HEADER
     //===============================================================================
     // SIEMENS AG / (c)Copyright 2021
     //-------------------------------------------------------------------------------
     // Title:            LStream_JsonSerializer
     // Comment/Function: parses a JSON string provided in the raw paramter
     //                   and rebuilds the coinatend bytes into a tree structure
     // Library/Family:   LStream
     // Author:           DI FA S SUP E&C
     // Tested with:      S7-1500 V2.8
     // Engineering:      TIA Portal V16
     // Restrictions:     -- 
     // Requirements:     LStream_typeElement(UDT)
     //-------------------------------------------------------------------------------
     // Change log table:
     // Version  | Date       | Expert in charge       | Changes applied
     //----------|------------|------------------------|------------------------------
     // 01.00.00 | 2021-06-10 | DI FA S SUP E&C        | First released version
     //===============================================================================
   END_REGION

   #tempExecute := #execute; // Work with temporary value / create process image

   REGION TRIGGERING
     IF (#tempExecute = TRUE) AND (#statExecuteOld = FALSE) // Check if FB is triggered
       AND (#statStatus = #STATUS_NO_CALL)
     THEN // First call; initialize FB
       #statDone := FALSE;
       #statBusy := TRUE;
       #statError := FALSE;
       #statStatus := #STATUS_FIRST_CALL;
       // State machine - start processing
       #statFbState := #FB_STATE_NEXT_ELEMENT;

       //Initialize functionality: reset OF variables, diagnostics, etc.
       #statJsonByteLen := UPPER_BOUND(ARR := #jsonByteArray, DIM := #FIRST_DIM);
       #statTreeLen := UPPER_BOUND(ARR := #tree, DIM := #FIRST_DIM);
       #statIndexTreeArray := 0;
       #statIndexJsonByteArray := 0;
       #statIsLastElement := FALSE;
       #statLastElementIsClosed := FALSE;
       #statStackIndex := -1;
       #statIsArrayOpen := FALSE;

     ELSIF (#statStatus = #STATUS_FIRST_CALL) THEN
       #statStatus := #STATUS_SUBSEQUENT_CALL;
     END_IF;

     // Edge detection 'execute' input
     #statExecuteOld := #tempExecute;
   END_REGION TRIGGERING

   IF (#statStatus = #STATUS_NO_CALL) THEN // Nothing to do -> End here to reduce "system load"
     RETURN;
   END_IF;

   REGION STATE_MACHINE

     //rest and start watchdog here so that repeat until has a maximum duration of constant MAX_LOOP_TIME
     #instWatchdog.TON(IN := FALSE,
                       PT := #MAX_REPEAT_TIME);
     //start watchdog
     #instWatchdog.TON(IN := TRUE,
                       PT := #MAX_REPEAT_TIME);
     REPEAT
       #statFbPreviousState := #statFbState;

       CASE #statFbState OF // State machine of FB

         #FB_STATE_NO_PROCESSING:
           REGION NO PROCESSING
             // No processing active (Note: this state must always be present and left empty)
             ;
           END_REGION NO PROCESSING

         #FB_STATE_NEXT_ELEMENT: // Work on next Element
           REGION NEXT_ELEMENT
             REGION ERROR HANDLING
               //check for last Element, either end of provided tree reached, or tree element is -1 = not initalized
               //this prevents index out of bounds error
               IF (#statIndexTreeArray = #statTreeLen - 1) OR #tree[#statIndexTreeArray + #NEXT_INDEX].type = #NOT_INITALYZED THEN
                 #statIsLastElement := TRUE;

               ELSIF (#statIndexTreeArray = #statTreeLen) THEN
                 //Error: Tree out of Bound
                 #statStatus := #ERR_TREE_OUT_OF_BOUNDS;
               END_IF;

               //Error: provided XML tree is too deep
               //max depth size allowed is size of stack, otherwise array out of bounds error will occur
               IF (#tree[#statIndexTreeArray].depth = #STACK_SIZE) THEN
                 #statStatus := #ERR_UNEXPECTED_DEPTH;
               ELSIF (#tree[#statIndexTreeArray].depth = #NOT_INITALYZED) THEN
                 //depth wasn't provided by user
                 #statStatus := #ERR_DEPTH_MISSING;
               END_IF;
             END_REGION #ERROR_HANDLING

             //must only be set once, reset after every new element
             #statIsFirstElement := FALSE;
             // stackIndex is used as current depth, is initalized wih -1 therefore first element, will always open an object 
             IF #statStackIndex < 0 THEN
               //open object
               #statInfoToWrite := CONCAT(IN1 := CHAR_TO_STRING(#BRACES_OPEN), IN2 := CHAR_TO_STRING(#WHITE_SPACE));
               //increase stack index and push closing elements on to it
               #statStackIndex += #INCREMENT_BY_ONE;
               #statStackIndexOpenElement[#statStackIndex] := #BRACES_CLOSE;
             END_IF;

             //in case Array is open, save the first key of the first field.
             //This is later used to check when new array field beginn 
             IF (#statIsArrayOpen AND #statFirstArrayKey = '') THEN

               //prevent that simple #ARRAY structure e.g "ArrayName":["ArrayValue1","ArrayValue2"]
               //is misread as key is array name that field info
               IF #statArrayName <> #tree[#statIndexTreeArray].key THEN
                 #statFirstArrayKey := #tree[#statIndexTreeArray].key;
               // ELSE //simple array case

               //   IF NOT #statIsFirstElement AND NOT #statIsSecondElement THEN
               //     //set flag that it is simple array
               //     //array field so no uneccarsy comma is written
               //     //as now depth change occurs
               //     #statIsFirstElement := TRUE;
               //   ELSE
               //     #statIsFirstElement := FALSE;
               //     #statIsSecondElement := TRUE;
               //   END_IF;
               END_IF;

               //in case Array is open, and current key matches first key of the first field,
               //indication of new array field, append open symbolic
             ELSIF (#statIsArrayOpen AND #statFirstArrayKey = #tree[#statIndexTreeArray].key) THEN

